   RUNG wire#w16
      Contact( "SMB_5" )
   END_RUNG wire#w17
   RUNG wire#w18
      Move(in := "MB_AD_RESET", out1 => "MB_DATA_MFC".MB_WRT_PARAM.DATA_ADDR)
      Move(in := 0, out1 => "MB_DATA_MFC".MB_WRT_PARAM.DATA_VAL)
   END_RUNG
   RUNG wire#powerrail
      Contact( #RUN )
      wire#w19
      Contact( "SMB_5" )
      Contact( "IEC_Timer_MFC_WRT_EVEN_DB".Q )
      wire#w20
      I_Contact( "SMB_7" )
      wire#w21
      Coil( "SMB_6" )
   END_RUNG
   RUNG wire#w19
      Contact( "SMB_6" )
   END_RUNG wire#w20
   RUNG wire#w21
      Move(in := "MB_VAL_RST_COUNTER", out1 => "MB_DATA_MFC".MB_WRT_PARAM.DATA_VAL)
   END_RUNG
   RUNG wire#powerrail
      Contact( #RUN )
      wire#w22
      Contact( "SMB_6" )
      Contact( "IEC_Timers_SMB_DB".Q )
      wire#w23
      I_Contact( "SMB_8" )
      wire#w24
      Coil( "SMB_7" )
   END_RUNG
   RUNG wire#w22
      Contact( "SMB_7" )
   END_RUNG wire#w23
   RUNG wire#w24
      Move(in := "MB_AD_COUNTER_MODE", out1 => "MB_DATA_MFC".MB_WRT_PARAM.DATA_ADDR)
      Move(in := "MB_VAL_COUNT_MODE_UP_LIMIT", out1 => "MB_DATA_MFC".MB_WRT_PARAM.DATA_VAL)
   END_RUNG
   RUNG wire#powerrail
      Contact( #RUN )
      wire#w25
      Contact( "SMB_7" )
      Contact( "IEC_Timer_MFC_WRT_EVEN_DB".Q )
      wire#w26
      Coil( "SMB_8" )
   END_RUNG
   RUNG wire#w25
      Contact( "SMB_8" )
   END_RUNG wire#w26
   RUNG wire#w26
      Coil( #ENDED )
   END_RUNG
   // the same network as SCL:
   #_w1 := #RUN AND #RUN AND NOT "SMB_M";   // rising edge of #RUN
   "SMB_M" := #RUN;
   "SMB_0" := (#_w1 OR (#RUN AND "SMB_0")) AND NOT "SMB_1" AND NOT "SMB_2";
   IF "SMB_0" THEN
       "MB_DATA_MFC".MB_WRT_PARAM.MB_ADDR := #MFC_ADDRESS;
       "MB_DATA_MFC".MB_WRT_PARAM.DATA_ADDR := "MB_AD_COUNTER_MODE";
       "MB_DATA_MFC".MB_WRT_PARAM.DATA_VAL := "MB_VAL_COUNT_MODE_OFF";
   END_IF;
   "SMB_1" := #RUN AND (("SMB_0" AND "IEC_Timers_SMB_DB".Q) OR "SMB_1") AND NOT "SMB_2" AND NOT "SMB_3";
   IF "SMB_1" THEN
       "MB_DATA_MFC".MB_WRT_PARAM.DATA_ADDR := "MB_AD_CONTROL_MODE";
       "MB_DATA_MFC".MB_WRT_PARAM.DATA_VAL := "MB_VAL_CONTROL_MODE_BUS";
   END_IF;
   "SMB_2" := #RUN AND (("SMB_1" AND "IEC_Timer_MFC_WRT_EVEN_DB".Q) OR "SMB_2") AND NOT "SMB_3" AND NOT "SMB_4";
   IF "SMB_2" THEN
       "MB_DATA_MFC".MB_WRT_PARAM.DATA_ADDR := "MB_AD_SETPOINT";
       "MB_DATA_MFC".MB_WRT_PARAM.DATA_VAL := #FLOW_SP;
   END_IF;
   "SMB_3" := #RUN AND (("SMB_2" AND "IEC_Timers_SMB_DB".Q) OR "SMB_3") AND NOT "SMB_4" AND NOT "SMB_5";
   IF "SMB_3" THEN
       "MB_DATA_MFC".MB_WRT_PARAM.DATA_ADDR := "MB_AD_COUNTER_LIMIT";
       "MB_DATA_MFC".MB_WRT_PARAM.DATA_VAL := #COUNTER_SP;
   END_IF;
   "SMB_4" := #RUN AND (("SMB_3" AND "IEC_Timer_MFC_WRT_EVEN_DB".Q) OR "SMB_4") AND NOT "SMB_5";
   IF "SMB_4" THEN
       "MB_DATA_MFC".MB_WRT_PARAM.DATA_ADDR := "MB_AD_COUNTER_SP_MODE";
       "MB_DATA_MFC".MB_WRT_PARAM.DATA_VAL := "MB_VAL_COUNT_SP_MODE_CHANGE";
   END_IF;
   "SMB_5" := #RUN AND (("SMB_4" AND "IEC_Timers_SMB_DB".Q) OR "SMB_5") AND NOT "SMB_6";
   IF "SMB_5" THEN
       "MB_DATA_MFC".MB_WRT_PARAM.DATA_ADDR := "MB_AD_RESET";
       "MB_DATA_MFC".MB_WRT_PARAM.DATA_VAL := 0;
   END_IF;
   "SMB_6" := #RUN AND (("SMB_5" AND "IEC_Timer_MFC_WRT_EVEN_DB".Q) OR "SMB_6") AND NOT "SMB_7";
   IF "SMB_6" THEN "MB_DATA_MFC".MB_WRT_PARAM.DATA_VAL := "MB_VAL_RST_COUNTER"; END_IF;
   "SMB_7" := #RUN AND (("SMB_6" AND "IEC_Timers_SMB_DB".Q) OR "SMB_7") AND NOT "SMB_8";
   IF "SMB_7" THEN
       "MB_DATA_MFC".MB_WRT_PARAM.DATA_ADDR := "MB_AD_COUNTER_MODE";
       "MB_DATA_MFC".MB_WRT_PARAM.DATA_VAL := "MB_VAL_COUNT_MODE_UP_LIMIT";
   END_IF;
   "SMB_8" := #RUN AND (("SMB_7" AND "IEC_Timer_MFC_WRT_EVEN_DB".Q) OR "SMB_8");
   #ENDED := "SMB_8";
END_REGION

REGION Network 2
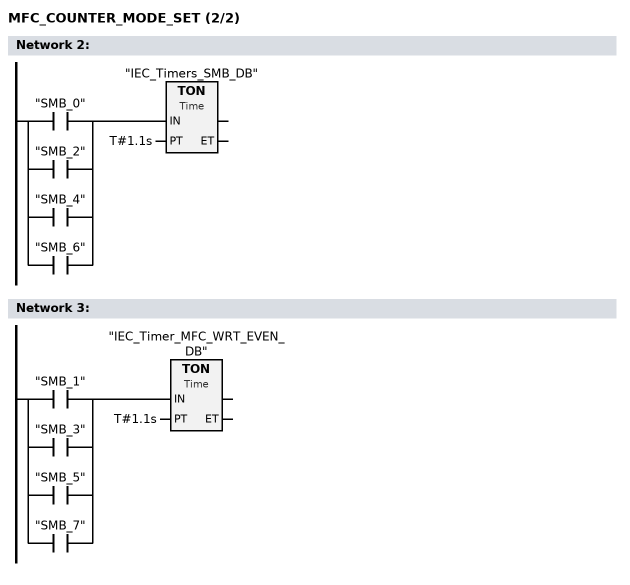
   "IEC_Timers_SMB_DB".TON(IN := "SMB_0" OR "SMB_2" OR "SMB_4" OR "SMB_6", PT := T#1.1s);
END_REGION

REGION Network 3
   "IEC_Timer_MFC_WRT_EVEN_DB".TON(IN := "SMB_1" OR "SMB_3" OR "SMB_5" OR "SMB_7", PT := T#1.1s);
END_REGION
END_FUNCTION

FUNCTION "ALL_VALVES_NORMAL" : Void   // FC20, LAD
{ S7_Optimized_Access := 'FALSE' }
VERSION : 0.1
BEGIN

REGION Network 1: NC
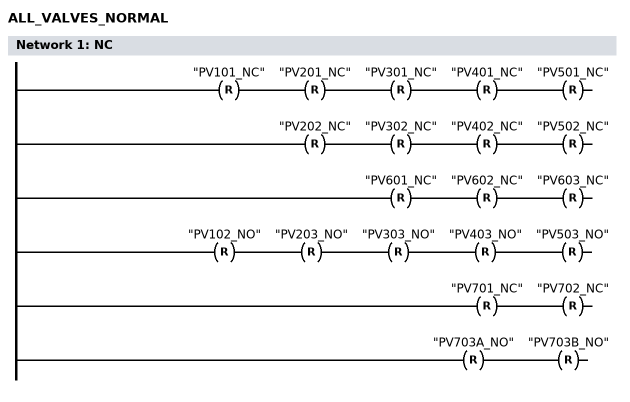
   RUNG wire#powerrail
      R_Coil( "PV101_NC" )
      R_Coil( "PV201_NC" )
      R_Coil( "PV301_NC" )
      R_Coil( "PV401_NC" )
      R_Coil( "PV501_NC" )
   END_RUNG
   RUNG wire#powerrail
      R_Coil( "PV202_NC" )
      R_Coil( "PV302_NC" )
      R_Coil( "PV402_NC" )
      R_Coil( "PV502_NC" )
   END_RUNG
   RUNG wire#powerrail
      R_Coil( "PV601_NC" )
      R_Coil( "PV602_NC" )
      R_Coil( "PV603_NC" )
   END_RUNG
   RUNG wire#powerrail
      R_Coil( "PV102_NO" )
      R_Coil( "PV203_NO" )
      R_Coil( "PV303_NO" )
      R_Coil( "PV403_NO" )
      R_Coil( "PV503_NO" )
   END_RUNG
   RUNG wire#powerrail
      R_Coil( "PV701_NC" )
      R_Coil( "PV702_NC" )
   END_RUNG
   RUNG wire#powerrail
      R_Coil( "PV703A_NO" )
      R_Coil( "PV703B_NO" )
   END_RUNG
   // the same network as SCL:
   "PV101_NC" := FALSE;
   "PV201_NC" := FALSE;
   "PV301_NC" := FALSE;
   "PV401_NC" := FALSE;
   "PV501_NC" := FALSE;
   "PV202_NC" := FALSE;
   "PV302_NC" := FALSE;
   "PV402_NC" := FALSE;
   "PV502_NC" := FALSE;
   "PV601_NC" := FALSE;
   "PV602_NC" := FALSE;
   "PV603_NC" := FALSE;
   "PV102_NO" := FALSE;
   "PV203_NO" := FALSE;
   "PV303_NO" := FALSE;
   "PV403_NO" := FALSE;
   "PV503_NO" := FALSE;
   "PV701_NC" := FALSE;
   "PV702_NC" := FALSE;
   "PV703A_NO" := FALSE;
   "PV703B_NO" := FALSE;
END_REGION
END_FUNCTION

FUNCTION "MFC_RESET" : Void   // FC21, LAD
{ S7_Optimized_Access := 'FALSE' }
VERSION : 0.1
   VAR_TEMP   // added for the SCL form of the ladder/FBD networks
      _w1 : Bool;
   END_VAR
BEGIN

REGION Network 1
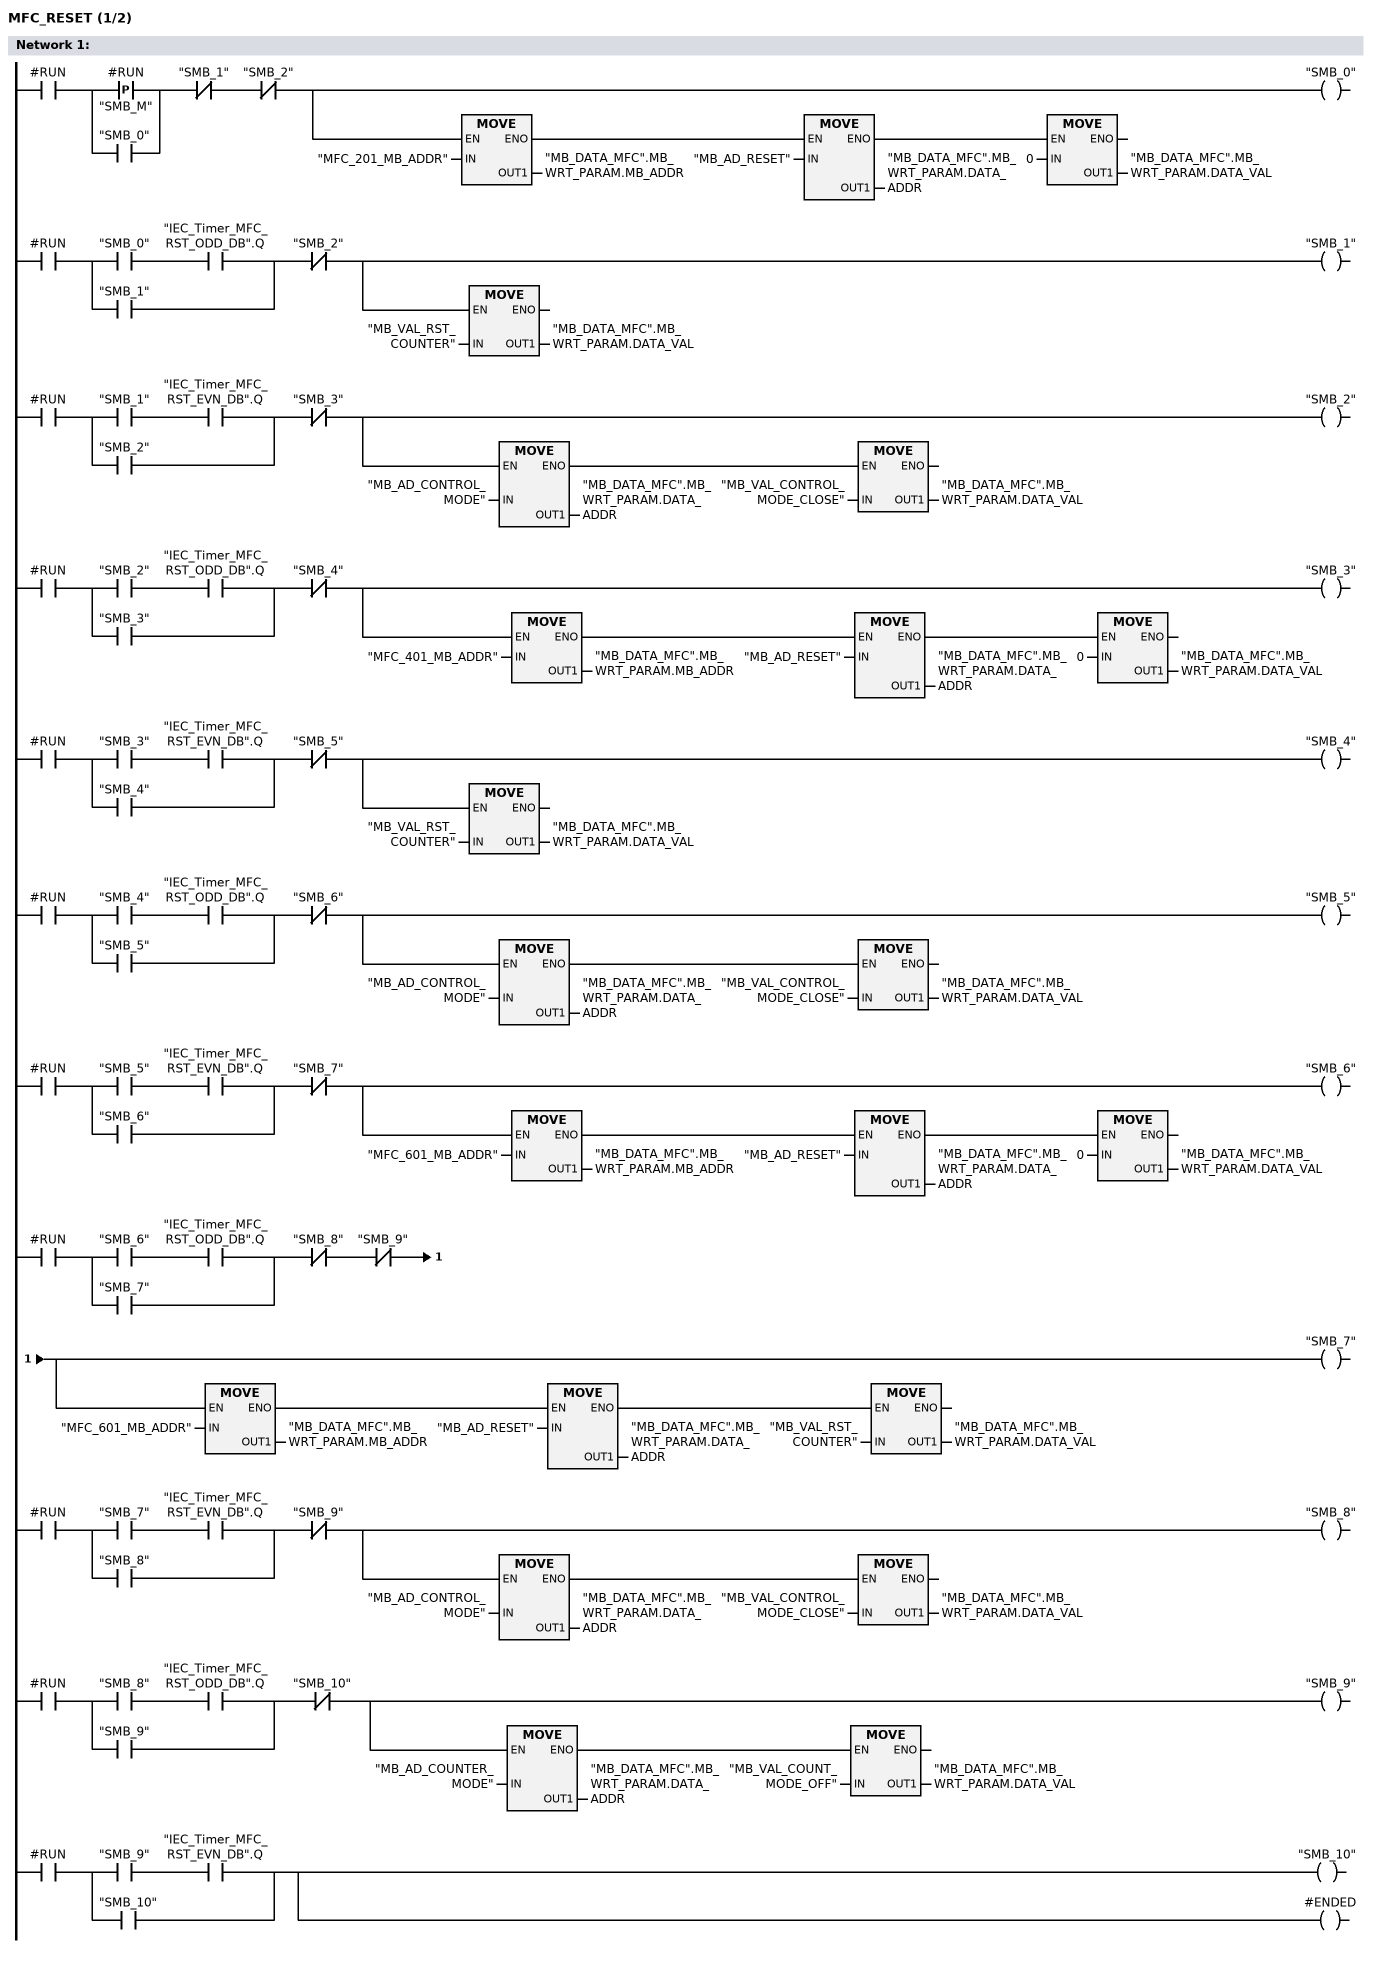
   RUNG wire#powerrail
      Contact( #RUN )
      wire#w1
      P_Contact(operand := #RUN, bit := "SMB_M")
      wire#w2
      I_Contact( "SMB_1" )
      I_Contact( "SMB_2" )
      wire#w3
      Coil( "SMB_0" )
   END_RUNG
   RUNG wire#w1
      Contact( "SMB_0" )
   END_RUNG wire#w2
   RUNG wire#w3
      Move(in := "MFC_201_MB_ADDR", out1 => "MB_DATA_MFC".MB_WRT_PARAM.MB_ADDR)
      Move(in := "MB_AD_RESET", out1 => "MB_DATA_MFC".MB_WRT_PARAM.DATA_ADDR)
      Move(in := 0, out1 => "MB_DATA_MFC".MB_WRT_PARAM.DATA_VAL)
   END_RUNG
   RUNG wire#powerrail
      Contact( #RUN )
      wire#w4
      Contact( "SMB_0" )
      Contact( "IEC_Timer_MFC_RST_ODD_DB".Q )
      wire#w5
      I_Contact( "SMB_2" )
      wire#w6
      Coil( "SMB_1" )
   END_RUNG
   RUNG wire#w4
      Contact( "SMB_1" )
   END_RUNG wire#w5
   RUNG wire#w6
      Move(in := "MB_VAL_RST_COUNTER", out1 => "MB_DATA_MFC".MB_WRT_PARAM.DATA_VAL)
   END_RUNG
   RUNG wire#powerrail
      Contact( #RUN )
      wire#w7
      Contact( "SMB_1" )
      Contact( "IEC_Timer_MFC_RST_EVN_DB".Q )
      wire#w8
      I_Contact( "SMB_3" )
      wire#w9
      Coil( "SMB_2" )
   END_RUNG
   RUNG wire#w7
      Contact( "SMB_2" )
   END_RUNG wire#w8
   RUNG wire#w9
      Move(in := "MB_AD_CONTROL_MODE", out1 => "MB_DATA_MFC".MB_WRT_PARAM.DATA_ADDR)
      Move(in := "MB_VAL_CONTROL_MODE_CLOSE", out1 => "MB_DATA_MFC".MB_WRT_PARAM.DATA_VAL)
   END_RUNG
   RUNG wire#powerrail
      Contact( #RUN )
      wire#w10
      Contact( "SMB_2" )
      Contact( "IEC_Timer_MFC_RST_ODD_DB".Q )
      wire#w11
      I_Contact( "SMB_4" )
      wire#w12
      Coil( "SMB_3" )
   END_RUNG
   RUNG wire#w10
      Contact( "SMB_3" )
   END_RUNG wire#w11
   RUNG wire#w12
      Move(in := "MFC_401_MB_ADDR", out1 => "MB_DATA_MFC".MB_WRT_PARAM.MB_ADDR)
      Move(in := "MB_AD_RESET", out1 => "MB_DATA_MFC".MB_WRT_PARAM.DATA_ADDR)
      Move(in := 0, out1 => "MB_DATA_MFC".MB_WRT_PARAM.DATA_VAL)
   END_RUNG
   RUNG wire#powerrail
      Contact( #RUN )
      wire#w13
      Contact( "SMB_3" )
      Contact( "IEC_Timer_MFC_RST_EVN_DB".Q )
      wire#w14
      I_Contact( "SMB_5" )
      wire#w15
      Coil( "SMB_4" )
   END_RUNG
   RUNG wire#w13
      Contact( "SMB_4" )
   END_RUNG wire#w14
   RUNG wire#w15
      Move(in := "MB_VAL_RST_COUNTER", out1 => "MB_DATA_MFC".MB_WRT_PARAM.DATA_VAL)
   END_RUNG
   RUNG wire#powerrail
      Contact( #RUN )
      wire#w16
      Contact( "SMB_4" )
      Contact( "IEC_Timer_MFC_RST_ODD_DB".Q )
      wire#w17
      I_Contact( "SMB_6" )
      wire#w18
      Coil( "SMB_5" )
   END_RUNG
   RUNG wire#w16
      Contact( "SMB_5" )
   END_RUNG wire#w17
   RUNG wire#w18
      Move(in := "MB_AD_CONTROL_MODE", out1 => "MB_DATA_MFC".MB_WRT_PARAM.DATA_ADDR)
      Move(in := "MB_VAL_CONTROL_MODE_CLOSE", out1 => "MB_DATA_MFC".MB_WRT_PARAM.DATA_VAL)
   END_RUNG
   RUNG wire#powerrail
      Contact( #RUN )
      wire#w19
      Contact( "SMB_5" )
      Contact( "IEC_Timer_MFC_RST_EVN_DB".Q )
      wire#w20
      I_Contact( "SMB_7" )
      wire#w21
      Coil( "SMB_6" )
   END_RUNG
   RUNG wire#w19
      Contact( "SMB_6" )
   END_RUNG wire#w20
   RUNG wire#w21
      Move(in := "MFC_601_MB_ADDR", out1 => "MB_DATA_MFC".MB_WRT_PARAM.MB_ADDR)
      Move(in := "MB_AD_RESET", out1 => "MB_DATA_MFC".MB_WRT_PARAM.DATA_ADDR)
      Move(in := 0, out1 => "MB_DATA_MFC".MB_WRT_PARAM.DATA_VAL)
   END_RUNG
   RUNG wire#powerrail
      Contact( #RUN )
      wire#w22
      Contact( "SMB_6" )
      Contact( "IEC_Timer_MFC_RST_ODD_DB".Q )
      wire#w23
      I_Contact( "SMB_8" )
      I_Contact( "SMB_9" )
      wire#w24
      Coil( "SMB_7" )
   END_RUNG
   RUNG wire#w22
      Contact( "SMB_7" )
   END_RUNG wire#w23
   RUNG wire#w24
      Move(in := "MFC_601_MB_ADDR", out1 => "MB_DATA_MFC".MB_WRT_PARAM.MB_ADDR)
      Move(in := "MB_AD_RESET", out1 => "MB_DATA_MFC".MB_WRT_PARAM.DATA_ADDR)
      Move(in := "MB_VAL_RST_COUNTER", out1 => "MB_DATA_MFC".MB_WRT_PARAM.DATA_VAL)
   END_RUNG
   RUNG wire#powerrail
      Contact( #RUN )
      wire#w25
      Contact( "SMB_7" )
      Contact( "IEC_Timer_MFC_RST_EVN_DB".Q )
      wire#w26
      I_Contact( "SMB_9" )
      wire#w27
      Coil( "SMB_8" )
   END_RUNG
   RUNG wire#w25
      Contact( "SMB_8" )
   END_RUNG wire#w26
   RUNG wire#w27
      Move(in := "MB_AD_CONTROL_MODE", out1 => "MB_DATA_MFC".MB_WRT_PARAM.DATA_ADDR)
      Move(in := "MB_VAL_CONTROL_MODE_CLOSE", out1 => "MB_DATA_MFC".MB_WRT_PARAM.DATA_VAL)
   END_RUNG
   RUNG wire#powerrail
      Contact( #RUN )
      wire#w28
      Contact( "SMB_8" )
      Contact( "IEC_Timer_MFC_RST_ODD_DB".Q )
      wire#w29
      I_Contact( "SMB_10" )
      wire#w30
      Coil( "SMB_9" )
   END_RUNG
   RUNG wire#w28
      Contact( "SMB_9" )
   END_RUNG wire#w29
   RUNG wire#w30
      Move(in := "MB_AD_COUNTER_MODE", out1 => "MB_DATA_MFC".MB_WRT_PARAM.DATA_ADDR)
      Move(in := "MB_VAL_COUNT_MODE_OFF", out1 => "MB_DATA_MFC".MB_WRT_PARAM.DATA_VAL)
   END_RUNG
   RUNG wire#powerrail
      Contact( #RUN )
      wire#w31
      Contact( "SMB_9" )
      Contact( "IEC_Timer_MFC_RST_EVN_DB".Q )
      wire#w32
      Coil( "SMB_10" )
   END_RUNG
   RUNG wire#w31
      Contact( "SMB_10" )
   END_RUNG wire#w32
   RUNG wire#w32
      Coil( #ENDED )
   END_RUNG
   // the same network as SCL:
   #_w1 := #RUN AND #RUN AND NOT "SMB_M";   // rising edge of #RUN
   "SMB_M" := #RUN;
   "SMB_0" := (#_w1 OR (#RUN AND "SMB_0")) AND NOT "SMB_1" AND NOT "SMB_2";
   IF "SMB_0" THEN
       "MB_DATA_MFC".MB_WRT_PARAM.MB_ADDR := "MFC_201_MB_ADDR";
       "MB_DATA_MFC".MB_WRT_PARAM.DATA_ADDR := "MB_AD_RESET";
       "MB_DATA_MFC".MB_WRT_PARAM.DATA_VAL := 0;
   END_IF;
   "SMB_1" := #RUN AND (("SMB_0" AND "IEC_Timer_MFC_RST_ODD_DB".Q) OR "SMB_1") AND NOT "SMB_2";
   IF "SMB_1" THEN "MB_DATA_MFC".MB_WRT_PARAM.DATA_VAL := "MB_VAL_RST_COUNTER"; END_IF;
   "SMB_2" := #RUN AND (("SMB_1" AND "IEC_Timer_MFC_RST_EVN_DB".Q) OR "SMB_2") AND NOT "SMB_3";
   IF "SMB_2" THEN
       "MB_DATA_MFC".MB_WRT_PARAM.DATA_ADDR := "MB_AD_CONTROL_MODE";
       "MB_DATA_MFC".MB_WRT_PARAM.DATA_VAL := "MB_VAL_CONTROL_MODE_CLOSE";
   END_IF;
   "SMB_3" := #RUN AND (("SMB_2" AND "IEC_Timer_MFC_RST_ODD_DB".Q) OR "SMB_3") AND NOT "SMB_4";
   IF "SMB_3" THEN
       "MB_DATA_MFC".MB_WRT_PARAM.MB_ADDR := "MFC_401_MB_ADDR";
       "MB_DATA_MFC".MB_WRT_PARAM.DATA_ADDR := "MB_AD_RESET";
       "MB_DATA_MFC".MB_WRT_PARAM.DATA_VAL := 0;
   END_IF;
   "SMB_4" := #RUN AND (("SMB_3" AND "IEC_Timer_MFC_RST_EVN_DB".Q) OR "SMB_4") AND NOT "SMB_5";
   IF "SMB_4" THEN "MB_DATA_MFC".MB_WRT_PARAM.DATA_VAL := "MB_VAL_RST_COUNTER"; END_IF;
   "SMB_5" := #RUN AND (("SMB_4" AND "IEC_Timer_MFC_RST_ODD_DB".Q) OR "SMB_5") AND NOT "SMB_6";
   IF "SMB_5" THEN
       "MB_DATA_MFC".MB_WRT_PARAM.DATA_ADDR := "MB_AD_CONTROL_MODE";
       "MB_DATA_MFC".MB_WRT_PARAM.DATA_VAL := "MB_VAL_CONTROL_MODE_CLOSE";
   END_IF;
   "SMB_6" := #RUN AND (("SMB_5" AND "IEC_Timer_MFC_RST_EVN_DB".Q) OR "SMB_6") AND NOT "SMB_7";
   IF "SMB_6" THEN
       "MB_DATA_MFC".MB_WRT_PARAM.MB_ADDR := "MFC_601_MB_ADDR";
       "MB_DATA_MFC".MB_WRT_PARAM.DATA_ADDR := "MB_AD_RESET";
       "MB_DATA_MFC".MB_WRT_PARAM.DATA_VAL := 0;
   END_IF;
   "SMB_7" := #RUN AND (("SMB_6" AND "IEC_Timer_MFC_RST_ODD_DB".Q) OR "SMB_7") AND NOT "SMB_8" AND NOT "SMB_9";
   IF "SMB_7" THEN
       "MB_DATA_MFC".MB_WRT_PARAM.MB_ADDR := "MFC_601_MB_ADDR";
       "MB_DATA_MFC".MB_WRT_PARAM.DATA_ADDR := "MB_AD_RESET";
       "MB_DATA_MFC".MB_WRT_PARAM.DATA_VAL := "MB_VAL_RST_COUNTER";
   END_IF;
   "SMB_8" := #RUN AND (("SMB_7" AND "IEC_Timer_MFC_RST_EVN_DB".Q) OR "SMB_8") AND NOT "SMB_9";
   IF "SMB_8" THEN
       "MB_DATA_MFC".MB_WRT_PARAM.DATA_ADDR := "MB_AD_CONTROL_MODE";
       "MB_DATA_MFC".MB_WRT_PARAM.DATA_VAL := "MB_VAL_CONTROL_MODE_CLOSE";
   END_IF;
   "SMB_9" := #RUN AND (("SMB_8" AND "IEC_Timer_MFC_RST_ODD_DB".Q) OR "SMB_9") AND NOT "SMB_10";
   IF "SMB_9" THEN
       "MB_DATA_MFC".MB_WRT_PARAM.DATA_ADDR := "MB_AD_COUNTER_MODE";
       "MB_DATA_MFC".MB_WRT_PARAM.DATA_VAL := "MB_VAL_COUNT_MODE_OFF";
   END_IF;
   "SMB_10" := #RUN AND (("SMB_9" AND "IEC_Timer_MFC_RST_EVN_DB".Q) OR "SMB_10");
   #ENDED := "SMB_10";
END_REGION

REGION Network 2
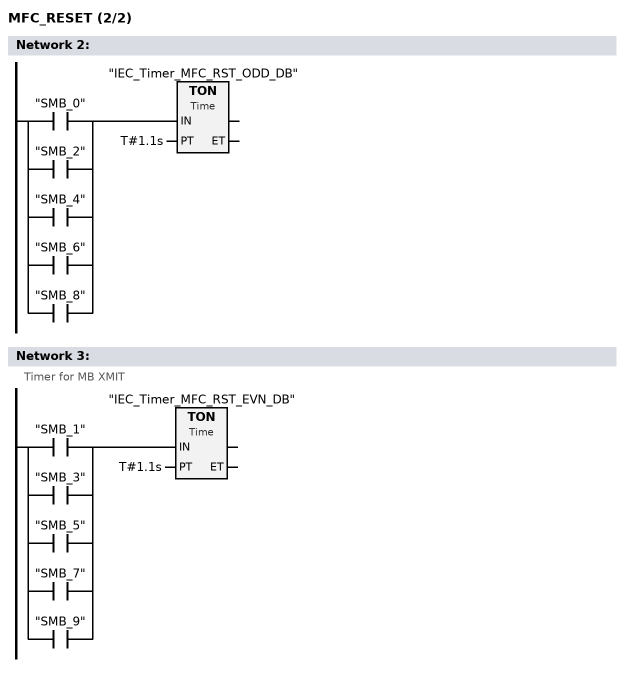
   "IEC_Timer_MFC_RST_ODD_DB".TON(IN := "SMB_0" OR "SMB_2" OR "SMB_4" OR "SMB_6" OR "SMB_8", PT := T#1.1s);
END_REGION

REGION Network 3
   // Timer for MB XMIT
   "IEC_Timer_MFC_RST_EVN_DB".TON(IN := "SMB_1" OR "SMB_3" OR "SMB_5" OR "SMB_7" OR "SMB_9", PT := T#1.1s);
END_REGION
END_FUNCTION

FUNCTION "ETAPA_1_HE_FC" : Void   // FC22, LAD
{ S7_Optimized_Access := 'FALSE' }
VERSION : 0.1
// Inertização da Câmara de testes com Helio. Max SP He =2.5 Bar
BEGIN

REGION Network 1: Alarm Set points
   // Alarm Set points of this step
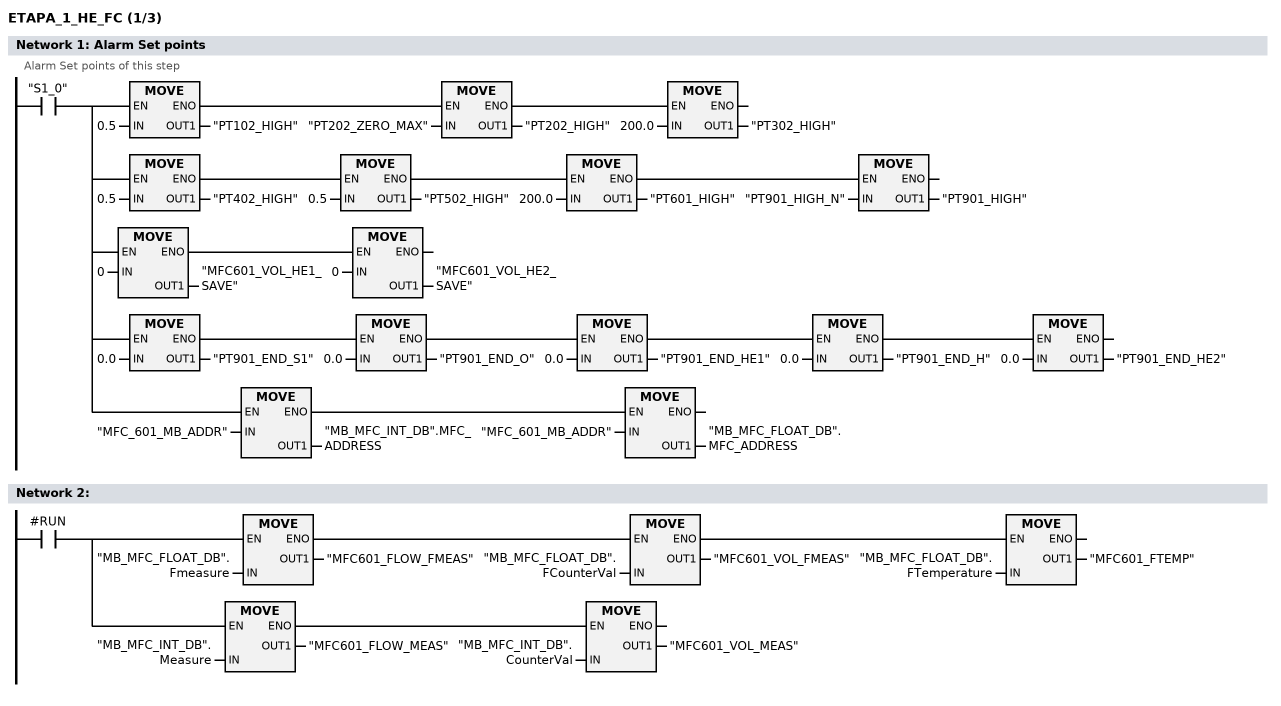
   RUNG wire#powerrail
      Contact( "S1_0" )
      wire#w1
      { S7_GenerateENO := "TRUE" } Move(in := 0.5, out1 => "PT102_HIGH")
      { S7_GenerateENO := "TRUE" } Move(in := "PT202_ZERO_MAX", out1 => "PT202_HIGH")
      { S7_GenerateENO := "TRUE" } Move(in := 200.0, out1 => "PT302_HIGH")
   END_RUNG
   RUNG wire#w1
      { S7_GenerateENO := "TRUE" } Move(in := 0.5, out1 => "PT402_HIGH")
      { S7_GenerateENO := "TRUE" } Move(in := 0.5, out1 => "PT502_HIGH")
      { S7_GenerateENO := "TRUE" } Move(in := 200.0, out1 => "PT601_HIGH")
      { S7_GenerateENO := "TRUE" } Move(in := "PT901_HIGH_N", out1 => "PT901_HIGH")
   END_RUNG
   RUNG wire#w1
      { S7_GenerateENO := "TRUE" } Move(in := 0, out1 => "MFC601_VOL_HE1_SAVE")
      { S7_GenerateENO := "TRUE" } Move(in := 0, out1 => "MFC601_VOL_HE2_SAVE")
   END_RUNG
   RUNG wire#w1
      { S7_GenerateENO := "TRUE" } Move(in := 0.0, out1 => "PT901_END_S1")
      { S7_GenerateENO := "TRUE" } Move(in := 0.0, out1 => "PT901_END_O")
      { S7_GenerateENO := "TRUE" } Move(in := 0.0, out1 => "PT901_END_HE1")
      { S7_GenerateENO := "TRUE" } Move(in := 0.0, out1 => "PT901_END_H")
      { S7_GenerateENO := "TRUE" } Move(in := 0.0, out1 => "PT901_END_HE2")
   END_RUNG
   RUNG wire#w1
      Move(in := "MFC_601_MB_ADDR", out1 => "MB_MFC_INT_DB".MFC_ADDRESS)
      Move(in := "MFC_601_MB_ADDR", out1 => "MB_MFC_FLOAT_DB".MFC_ADDRESS)
   END_RUNG
   // the same network as SCL:
   // ENO of a box is taken as its EN; it also drops when the box reports an error
   IF "S1_0" THEN
       "PT102_HIGH" := 0.5;
       "PT202_HIGH" := "PT202_ZERO_MAX";
       "PT302_HIGH" := 200.0;
       "PT402_HIGH" := 0.5;
       "PT502_HIGH" := 0.5;
       "PT601_HIGH" := 200.0;
       "PT901_HIGH" := "PT901_HIGH_N";
       "MFC601_VOL_HE1_SAVE" := 0;
       "MFC601_VOL_HE2_SAVE" := 0;
       "PT901_END_S1" := 0.0;
       "PT901_END_O" := 0.0;
       "PT901_END_HE1" := 0.0;
       "PT901_END_H" := 0.0;
       "PT901_END_HE2" := 0.0;
       "MB_MFC_INT_DB".MFC_ADDRESS := "MFC_601_MB_ADDR";
       "MB_MFC_FLOAT_DB".MFC_ADDRESS := "MFC_601_MB_ADDR";
   END_IF;
END_REGION

REGION Network 2
   RUNG wire#powerrail
      Contact( #RUN )
      wire#w1
      { S7_GenerateENO := "TRUE" } Move(in := "MB_MFC_FLOAT_DB".Fmeasure, out1 => "MFC601_FLOW_FMEAS")
      { S7_GenerateENO := "TRUE" } Move(in := "MB_MFC_FLOAT_DB".FCounterVal, out1 => "MFC601_VOL_FMEAS")
      { S7_GenerateENO := "TRUE" } Move(in := "MB_MFC_FLOAT_DB".FTemperature, out1 => "MFC601_FTEMP")
   END_RUNG
   RUNG wire#w1
      { S7_GenerateENO := "TRUE" } Move(in := "MB_MFC_INT_DB".Measure, out1 => "MFC601_FLOW_MEAS")
      { S7_GenerateENO := "TRUE" } Move(in := "MB_MFC_INT_DB".CounterVal, out1 => "MFC601_VOL_MEAS")
   END_RUNG
   // the same network as SCL:
   // ENO of a box is taken as its EN; it also drops when the box reports an error
   IF #RUN THEN
       "MFC601_FLOW_FMEAS" := "MB_MFC_FLOAT_DB".Fmeasure;
       "MFC601_VOL_FMEAS" := "MB_MFC_FLOAT_DB".FCounterVal;
       "MFC601_FTEMP" := "MB_MFC_FLOAT_DB".FTemperature;
       "MFC601_FLOW_MEAS" := "MB_MFC_INT_DB".Measure;
       "MFC601_VOL_MEAS" := "MB_MFC_INT_DB".CounterVal;
   END_IF;
END_REGION

REGION Network 3
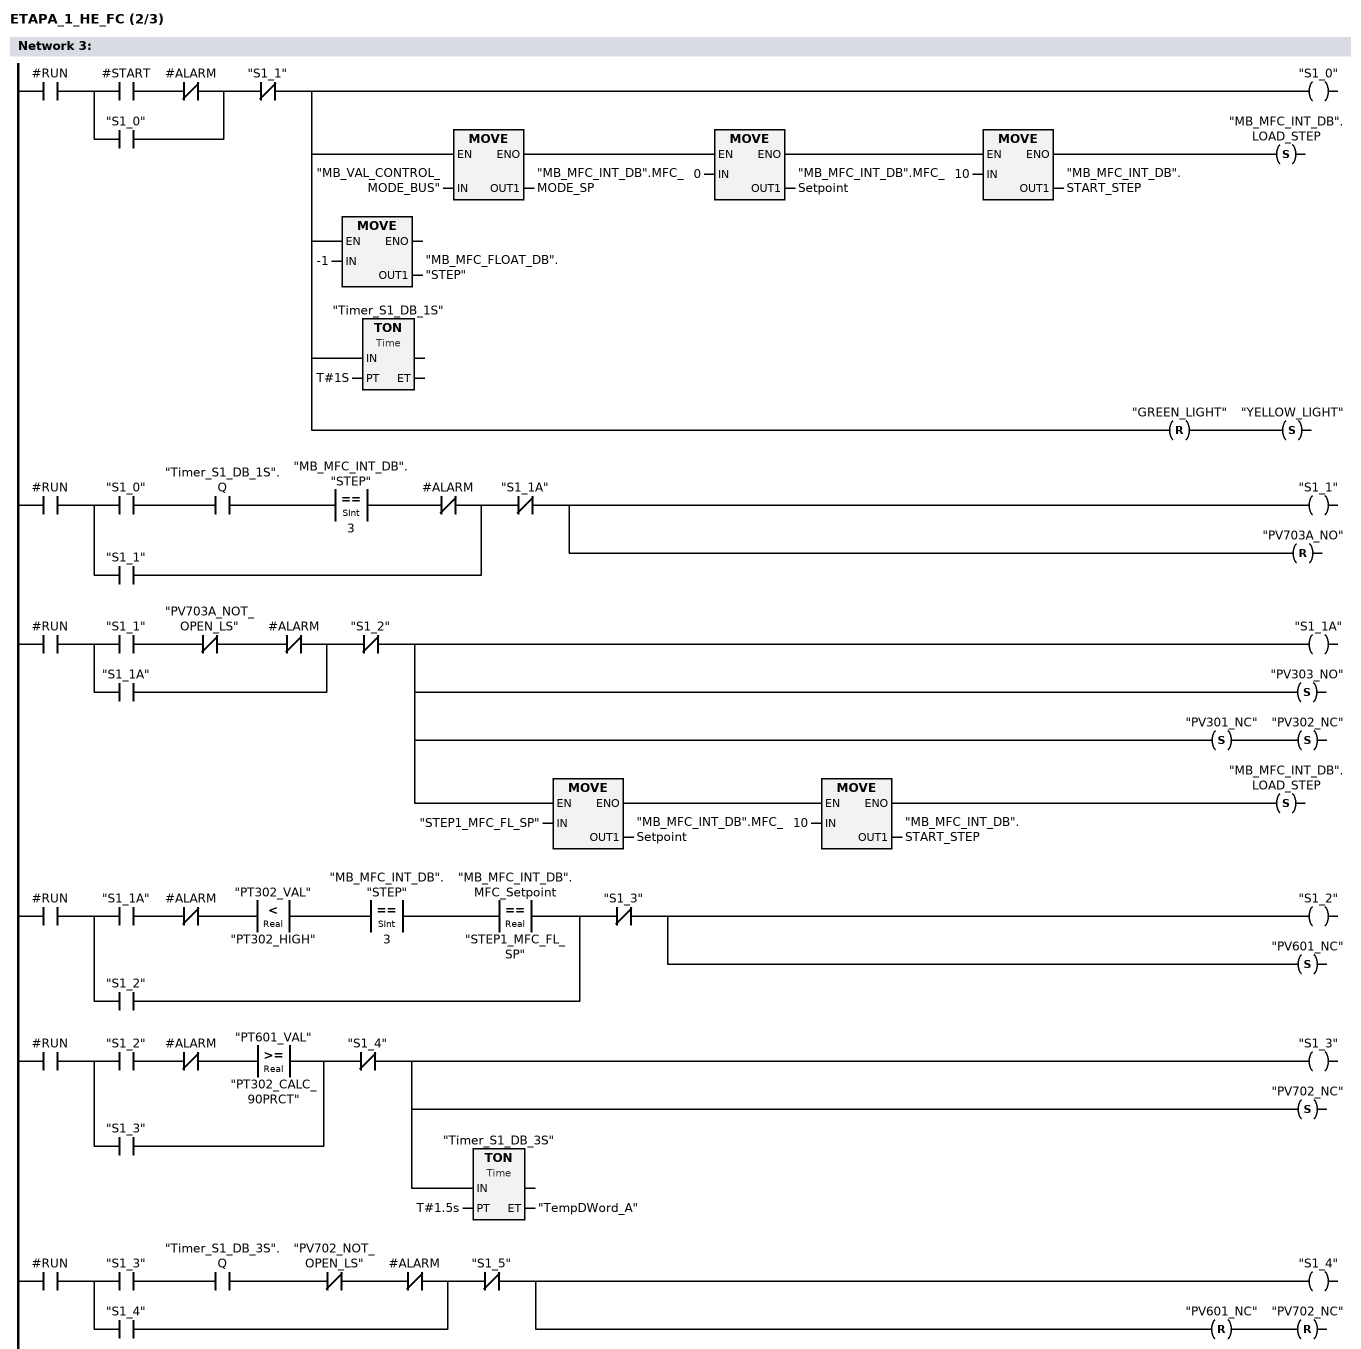
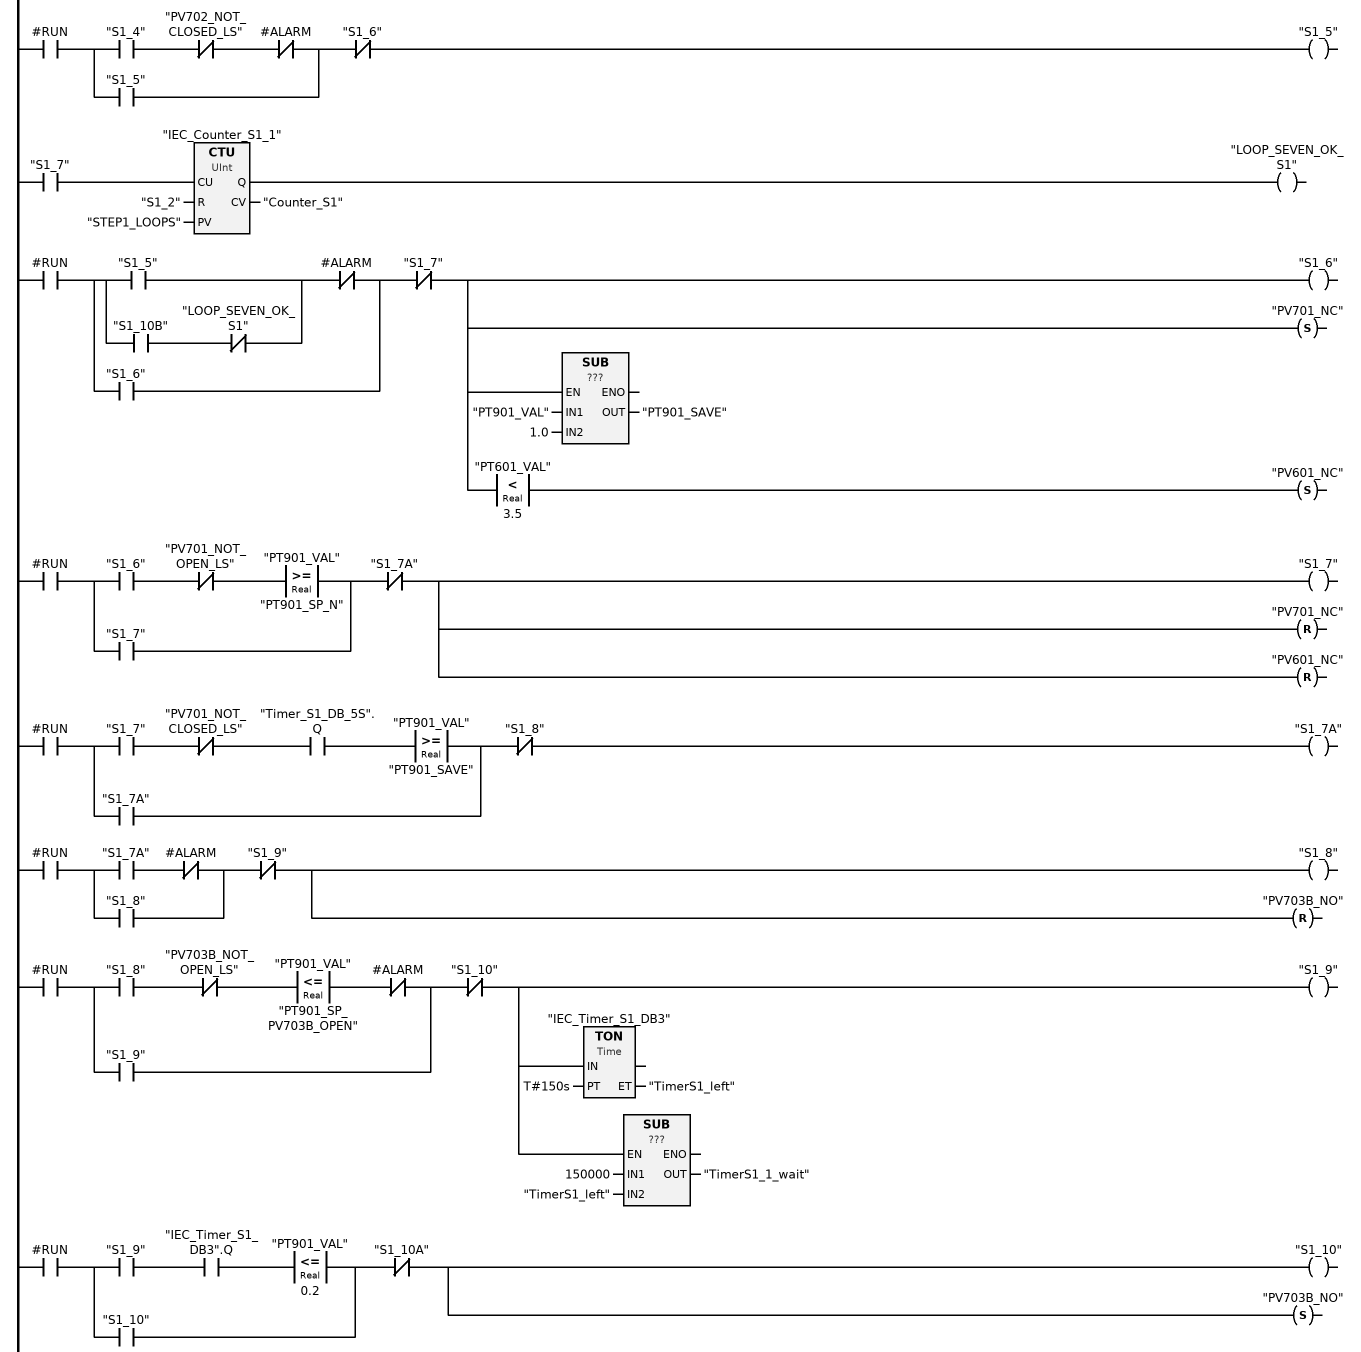